REGION Network 6: setare bit 1 pentru SERVO6
   RUNG wire#powerrail
      I_Contact( "DB_HMI"."MAN/AUTO" )
      Contact( "DB_HMI_buttons"."ON/OFF_servo6" )
      wire#w1
      S_SR(operand := "DB_06_Write_Arduino".Servo6, r1 := wire#w3)
   END_RUNG
   RUNG wire#powerrail
      Contact( "DB_HMI"."MAN/AUTO" )
      Contact( "DB_Markers_Auto".servo6_auto )
   END_RUNG wire#w1
   RUNG wire#powerrail
      I_Contact( "DB_HMI"."MAN/AUTO" )
      I_Contact( "DB_HMI_buttons"."ON/OFF_servo6" )
      wire#w2
      R_Coil( "DB_HMI_buttons"."ON/OFF_servo6" )
   END_RUNG wire#w3
   RUNG wire#powerrail
      Contact( "DB_HMI"."MAN/AUTO" )
      I_Contact( "DB_Markers_Auto".servo6_auto )
   END_RUNG wire#w2
   RUNG wire#powerrail
      Contact( "DB_HMI_buttons".STOP )
   END_RUNG wire#w2
   // the same network as SCL:
   #_w1 := (NOT "DB_HMI"."MAN/AUTO" AND NOT "DB_HMI_buttons"."ON/OFF_servo6") OR ("DB_HMI"."MAN/AUTO" AND NOT "DB_Markers_Auto".servo6_auto) OR "DB_HMI_buttons".STOP;
   #_w2 := (NOT "DB_HMI"."MAN/AUTO" AND "DB_HMI_buttons"."ON/OFF_servo6") OR ("DB_HMI"."MAN/AUTO" AND "DB_Markers_Auto".servo6_auto);
   IF #_w1 THEN "DB_HMI_buttons"."ON/OFF_servo6" := FALSE; END_IF;
   IF #_w2 THEN
       "DB_06_Write_Arduino".Servo6 := TRUE;   // SR flip-flop
   END_IF;
   IF #_w1 THEN "DB_06_Write_Arduino".Servo6 := FALSE; END_IF;
END_REGION

REGION Network 7: setare bit stepper2_up
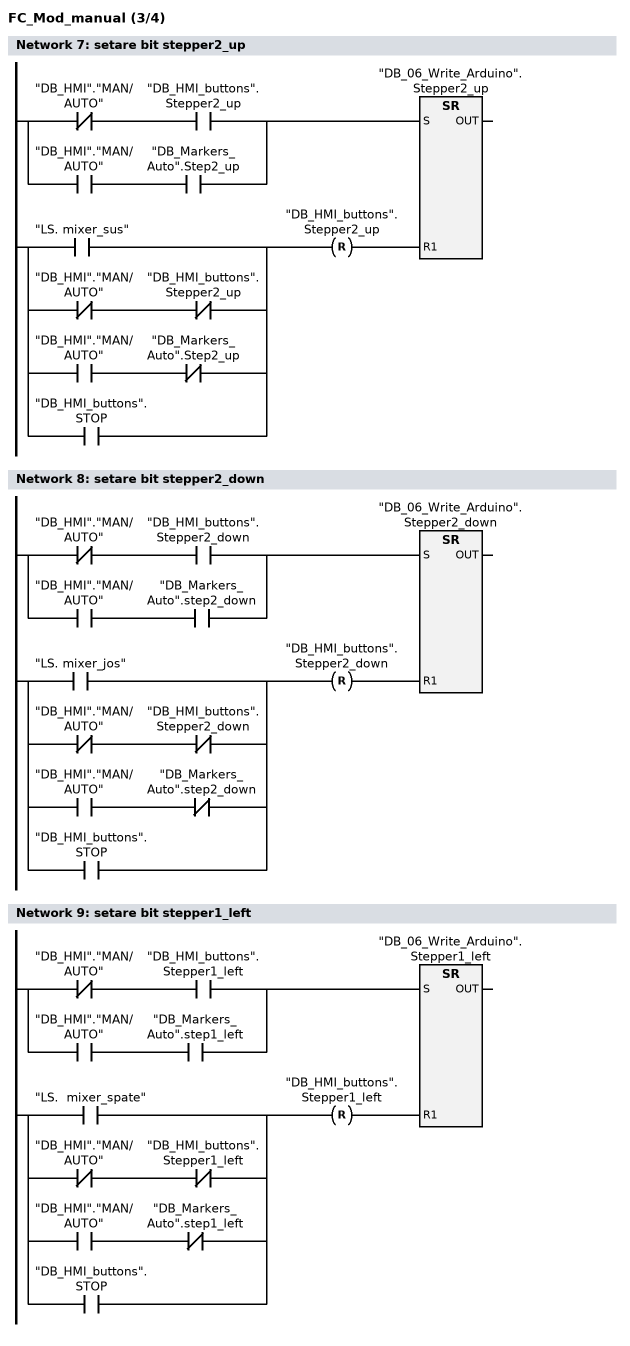
   RUNG wire#powerrail
      I_Contact( "DB_HMI"."MAN/AUTO" )
      Contact( "DB_HMI_buttons".Stepper2_up )
      wire#w1
      S_SR(operand := "DB_06_Write_Arduino".Stepper2_up, r1 := wire#w3)
   END_RUNG
   RUNG wire#powerrail
      Contact( "DB_HMI"."MAN/AUTO" )
      Contact( "DB_Markers_Auto".Step2_up )
   END_RUNG wire#w1
   RUNG wire#powerrail
      Contact( "LS. mixer_sus" )
      wire#w2
      R_Coil( "DB_HMI_buttons".Stepper2_up )
   END_RUNG wire#w3
   RUNG wire#powerrail
      I_Contact( "DB_HMI"."MAN/AUTO" )
      I_Contact( "DB_HMI_buttons".Stepper2_up )
   END_RUNG wire#w2
   RUNG wire#powerrail
      Contact( "DB_HMI"."MAN/AUTO" )
      I_Contact( "DB_Markers_Auto".Step2_up )
   END_RUNG wire#w2
   RUNG wire#powerrail
      Contact( "DB_HMI_buttons".STOP )
   END_RUNG wire#w2
   // the same network as SCL:
   #_w1 := "LS. mixer_sus" OR (NOT "DB_HMI"."MAN/AUTO" AND NOT "DB_HMI_buttons".Stepper2_up) OR ("DB_HMI"."MAN/AUTO" AND NOT "DB_Markers_Auto".Step2_up) OR "DB_HMI_buttons".STOP;
   #_w2 := (NOT "DB_HMI"."MAN/AUTO" AND "DB_HMI_buttons".Stepper2_up) OR ("DB_HMI"."MAN/AUTO" AND "DB_Markers_Auto".Step2_up);
   IF #_w1 THEN "DB_HMI_buttons".Stepper2_up := FALSE; END_IF;
   IF #_w2 THEN
       "DB_06_Write_Arduino".Stepper2_up := TRUE;   // SR flip-flop
   END_IF;
   IF #_w1 THEN "DB_06_Write_Arduino".Stepper2_up := FALSE; END_IF;
END_REGION

REGION Network 8: setare bit stepper2_down
   RUNG wire#powerrail
      I_Contact( "DB_HMI"."MAN/AUTO" )
      Contact( "DB_HMI_buttons".Stepper2_down )
      wire#w1
      S_SR(operand := "DB_06_Write_Arduino".Stepper2_down, r1 := wire#w3)
   END_RUNG
   RUNG wire#powerrail
      Contact( "DB_HMI"."MAN/AUTO" )
      Contact( "DB_Markers_Auto".step2_down )
   END_RUNG wire#w1
   RUNG wire#powerrail
      Contact( "LS. mixer_jos" )
      wire#w2
      R_Coil( "DB_HMI_buttons".Stepper2_down )
   END_RUNG wire#w3
   RUNG wire#powerrail
      I_Contact( "DB_HMI"."MAN/AUTO" )
      I_Contact( "DB_HMI_buttons".Stepper2_down )
   END_RUNG wire#w2
   RUNG wire#powerrail
      Contact( "DB_HMI"."MAN/AUTO" )
      I_Contact( "DB_Markers_Auto".step2_down )
   END_RUNG wire#w2
   RUNG wire#powerrail
      Contact( "DB_HMI_buttons".STOP )
   END_RUNG wire#w2
   // the same network as SCL:
   #_w1 := "LS. mixer_jos" OR (NOT "DB_HMI"."MAN/AUTO" AND NOT "DB_HMI_buttons".Stepper2_down) OR ("DB_HMI"."MAN/AUTO" AND NOT "DB_Markers_Auto".step2_down) OR "DB_HMI_buttons".STOP;
   #_w2 := (NOT "DB_HMI"."MAN/AUTO" AND "DB_HMI_buttons".Stepper2_down) OR ("DB_HMI"."MAN/AUTO" AND "DB_Markers_Auto".step2_down);
   IF #_w1 THEN "DB_HMI_buttons".Stepper2_down := FALSE; END_IF;
   IF #_w2 THEN
       "DB_06_Write_Arduino".Stepper2_down := TRUE;   // SR flip-flop
   END_IF;
   IF #_w1 THEN "DB_06_Write_Arduino".Stepper2_down := FALSE; END_IF;
END_REGION

REGION Network 9: setare bit stepper1_left
   RUNG wire#powerrail
      I_Contact( "DB_HMI"."MAN/AUTO" )
      Contact( "DB_HMI_buttons".Stepper1_left )
      wire#w1
      S_SR(operand := "DB_06_Write_Arduino".Stepper1_left, r1 := wire#w3)
   END_RUNG
   RUNG wire#powerrail
      Contact( "DB_HMI"."MAN/AUTO" )
      Contact( "DB_Markers_Auto".step1_left )
   END_RUNG wire#w1
   RUNG wire#powerrail
      Contact( "LS.  mixer_spate" )
      wire#w2
      R_Coil( "DB_HMI_buttons".Stepper1_left )
   END_RUNG wire#w3
   RUNG wire#powerrail
      I_Contact( "DB_HMI"."MAN/AUTO" )
      I_Contact( "DB_HMI_buttons".Stepper1_left )
   END_RUNG wire#w2
   RUNG wire#powerrail
      Contact( "DB_HMI"."MAN/AUTO" )
      I_Contact( "DB_Markers_Auto".step1_left )
   END_RUNG wire#w2
   RUNG wire#powerrail
      Contact( "DB_HMI_buttons".STOP )
   END_RUNG wire#w2
   // the same network as SCL:
   #_w1 := "LS.  mixer_spate" OR (NOT "DB_HMI"."MAN/AUTO" AND NOT "DB_HMI_buttons".Stepper1_left) OR ("DB_HMI"."MAN/AUTO" AND NOT "DB_Markers_Auto".step1_left) OR "DB_HMI_buttons".STOP;
   #_w2 := (NOT "DB_HMI"."MAN/AUTO" AND "DB_HMI_buttons".Stepper1_left) OR ("DB_HMI"."MAN/AUTO" AND "DB_Markers_Auto".step1_left);
   IF #_w1 THEN "DB_HMI_buttons".Stepper1_left := FALSE; END_IF;
   IF #_w2 THEN
       "DB_06_Write_Arduino".Stepper1_left := TRUE;   // SR flip-flop
   END_IF;
   IF #_w1 THEN "DB_06_Write_Arduino".Stepper1_left := FALSE; END_IF;
END_REGION

REGION Network 10: setare bit stepper1_right
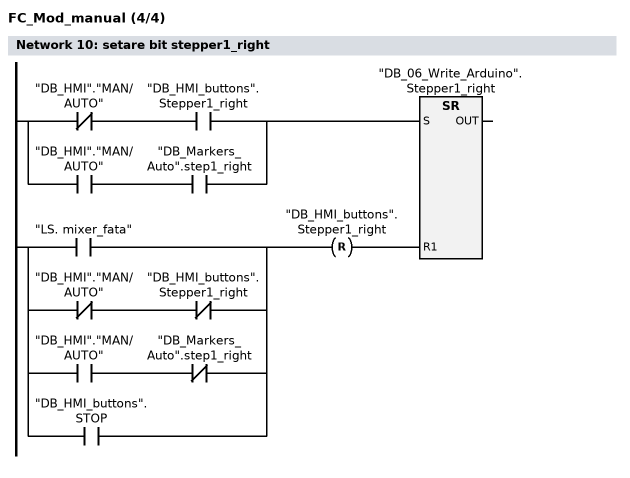
   RUNG wire#powerrail
      I_Contact( "DB_HMI"."MAN/AUTO" )
      Contact( "DB_HMI_buttons".Stepper1_right )
      wire#w1
      S_SR(operand := "DB_06_Write_Arduino".Stepper1_right, r1 := wire#w3)
   END_RUNG
   RUNG wire#powerrail
      Contact( "DB_HMI"."MAN/AUTO" )
      Contact( "DB_Markers_Auto".step1_right )
   END_RUNG wire#w1
   RUNG wire#powerrail
      Contact( "LS. mixer_fata" )
      wire#w2
      R_Coil( "DB_HMI_buttons".Stepper1_right )
   END_RUNG wire#w3
   RUNG wire#powerrail
      I_Contact( "DB_HMI"."MAN/AUTO" )
      I_Contact( "DB_HMI_buttons".Stepper1_right )
   END_RUNG wire#w2
   RUNG wire#powerrail
      Contact( "DB_HMI"."MAN/AUTO" )
      I_Contact( "DB_Markers_Auto".step1_right )
   END_RUNG wire#w2
   RUNG wire#powerrail
      Contact( "DB_HMI_buttons".STOP )
   END_RUNG wire#w2
   // the same network as SCL:
   #_w1 := "LS. mixer_fata" OR (NOT "DB_HMI"."MAN/AUTO" AND NOT "DB_HMI_buttons".Stepper1_right) OR ("DB_HMI"."MAN/AUTO" AND NOT "DB_Markers_Auto".step1_right) OR "DB_HMI_buttons".STOP;
   #_w2 := (NOT "DB_HMI"."MAN/AUTO" AND "DB_HMI_buttons".Stepper1_right) OR ("DB_HMI"."MAN/AUTO" AND "DB_Markers_Auto".step1_right);
   IF #_w1 THEN "DB_HMI_buttons".Stepper1_right := FALSE; END_IF;
   IF #_w2 THEN
       "DB_06_Write_Arduino".Stepper1_right := TRUE;   // SR flip-flop
   END_IF;
   IF #_w1 THEN "DB_06_Write_Arduino".Stepper1_right := FALSE; END_IF;
END_REGION
END_FUNCTION

FUNCTION "FC_select_reteta_FBD_language" : Void   // FC8, FBD
{ S7_Optimized_Access := 'TRUE' }
VERSION : 0.1
BEGIN

REGION Network 1: Reteta ciocolata neagra =1
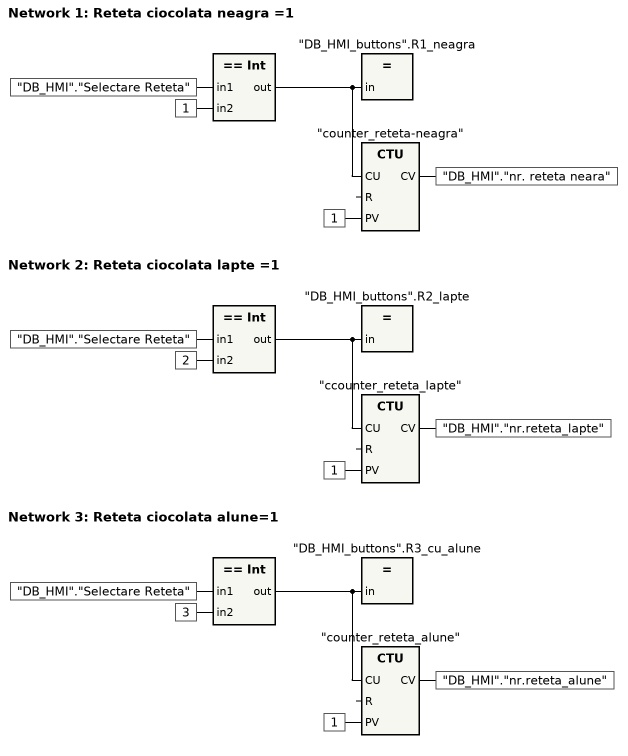
   "DB_HMI_buttons".R1_neagra := "DB_HMI"."Selectare Reteta" = 1;
   "counter_reteta-neagra".CTU(CU := "DB_HMI_buttons".R1_neagra, PV := 1, CV => "DB_HMI"."nr. reteta neara");
END_REGION

REGION Network 2: Reteta ciocolata lapte =1
   "DB_HMI_buttons".R2_lapte := "DB_HMI"."Selectare Reteta" = 2;
   "ccounter_reteta_lapte".CTU(CU := "DB_HMI_buttons".R2_lapte, PV := 1, CV => "DB_HMI"."nr.reteta_lapte");
END_REGION

REGION Network 3: Reteta ciocolata alune=1
   "DB_HMI_buttons".R3_cu_alune := "DB_HMI"."Selectare Reteta" = 3;
   "counter_reteta_alune".CTU(CU := "DB_HMI_buttons".R3_cu_alune, PV := 1, CV => "DB_HMI"."nr.reteta_alune");
END_REGION
END_FUNCTION

(* ===== HMI "HMI_RT_1" =====
system functions are stored by id; their names below are inferred from use
connection "Connection_1": ETHERNET, SMART_S7_1500_OMS
connection "HMI_Connection_1": ETHERNET, SMART_S7_1500_OMS

HMI tags "Default tag table"
   "LS_left" : Bool = PLC "LS.  mixer_spate" AT %I10.5, 1 s
   "LS_right" : Bool = PLC "LS. mixer_fata" AT %I10.2, 1 s
   "LS_up" : Bool = PLC "LS. mixer_sus" AT %I10.6, 1 s
   "LS_down" : Bool = PLC "LS. mixer_jos" AT %I10.1, 1 s
   "DB_HMI_BUTTON_DEV1:PLITA" : Bool = PLC DB_HMI_buttons.ON/OFF_plita AT %DB1.DBX0.0, 1 s
   "DB_HMI_BUTTON_DEV2:Mixer" : Bool = PLC DB_HMI_buttons.ON/OFF_mixer AT %DB1.DBX0.0, 1 s
   "DB_HMI_BUTTON_DEV2:Pompa" : Bool = PLC DB_HMI_buttons.ON/OFF_pompa AT %DB1.DBX0.0, 1 s
   "Reset ciuperca" : Bool = PLC DB_HMI_buttons.Reset_ciuperca AT %DB1.DBX0.0, 1 s
   "DB_06_Write_Arduino_Servo1" : Bool = PLC DB_06_Write_Arduino.Servo1 AT %DB6.DBX0.0, 1 s
   "DB_06_Write_Arduino_Servo2" : Bool = PLC DB_06_Write_Arduino.Servo2 AT %DB6.DBX0.1, 1 s
   "DB_06_Write_Arduino_Servo3" : Bool = PLC DB_06_Write_Arduino.Servo3 AT %DB6.DBX0.2, 1 s
   "DB_06_Write_Arduino_Servo4" : Bool = PLC DB_06_Write_Arduino.Servo4 AT %DB6.DBX0.3, 1 s
   "DB_06_Write_Arduino_Servo5" : Bool = PLC DB_06_Write_Arduino.Servo5 AT %DB6.DBX0.4, 1 s
   "DB_06_Write_Arduino_Servo6" : Bool = PLC DB_06_Write_Arduino.Servo6 AT %DB6.DBX0.5, 1 s
   "DB_HMI_buttons_ON/OFF_servo1" : Bool = PLC DB_HMI_buttons.ON/OFF_servo1, 1 s
   "ON/OFF_Servo1_HMI" : Word = PLC "ON/OFF_Servo1_HMI" AT %MW2, 1 s
   "ON/OFF_servo2_HMI" : Word = PLC "ON/OFF_servo2_HMI" AT %MW4, 1 s
   "ON/OFF_SERVO3_HMI" : Word = PLC "ON/OFF_SERVO3_HMI" AT %MW6, 1 s
   "ON/OFF_SERVO4_HMI" : Word = PLC "ON/OFF_SERVO4_HMI" AT %MW14, 1 s
   "ON/OFF_SERVO5_HMI" : Word = PLC "ON/OFF_SERVO5_HMI" AT %MW16, 1 s
   "ON/OFF_SERVO6_HMI" : Word = PLC "ON/OFF_SERVO6_HMI" AT %MW18, 1 s
   "ON/OFF_servo1" : Bool = PLC "ON/OFF_servo1" AT %M1.4, 1 s
   "DB_HMI_buttons_ON/OFF_servo2" : Bool = PLC DB_HMI_buttons.ON/OFF_servo2, 1 s
   "DB_HMI_buttons_ON/OFF_servo3" : Bool = PLC DB_HMI_buttons.ON/OFF_servo3, 1 s
   "DB_HMI_buttons_ON/OFF_servo4" : Bool = PLC DB_HMI_buttons.ON/OFF_servo4, 1 s
   "DB_HMI_buttons_ON/OFF_servo5" : Bool = PLC DB_HMI_buttons.ON/OFF_servo5, 1 s
   "DB_HMI_buttons_ON/OFF_servo6" : Bool = PLC DB_HMI_buttons.ON/OFF_servo6, 1 s
   "DB_HMI_buttons_Reset" : Bool = PLC DB_HMI_buttons.Reset, 1 s
   "DB_HMI_buttons_STOP" : Bool = PLC DB_HMI_buttons.STOP, 1 s
   "Reteta" : Int = PLC DB_HMI_buttons.Reteta_text_list AT %DB1.DBX0.0, 1 s
   "Start_initializare" : Bool = PLC DB_HMI_buttons.Start/Stop_initializare, 1 s
   "Start_proces" : Bool = PLC DB_HMI_buttons.Start/Stop_proces_auto, 1 s
   "DB_03_Read_Arduino_temp_citita" : Real = PLC DB_03_Read_Arduino.temp_citita AT %DB3.DBD0, 1 s
   "DB_06_Write_Arduino_Stepper2_up" : Bool = PLC DB_06_Write_Arduino.Stepper2_up AT %DB6.DBX1.0, 1 s
   "DB_06_Write_Arduino_Stepper2_down" : Bool = PLC DB_06_Write_Arduino.Stepper2_down AT %DB6.DBX1.1, 1 s
   "DB_HMI_buttons_Curatare" : Bool = PLC DB_HMI_buttons.Curatare, 1 s
   "DB_HMI_MAN/AUTO" : Bool = PLC DB_HMI.MAN/AUTO, 1 s
   "DB_HMI_Selectare Reteta" : Int = PLC DB_HMI."Selectare Reteta", 1 s
   "DB_06_Write_Arduino_Stepper1_left" : Bool = PLC DB_06_Write_Arduino.Stepper1_left AT %DB6.DBX0.6, 1 s
   "DB_06_Write_Arduino_Stepper1_right" : Bool = PLC DB_06_Write_Arduino.Stepper1_right AT %DB6.DBX0.7, 1 s
   "DB_HMI_buttons_Stepper1_left" : Bool = PLC DB_HMI_buttons.Stepper1_left, 1 s
   "DB_HMI_buttons_Stepper1_right" : Bool = PLC DB_HMI_buttons.Stepper1_right, 1 s
   "DB_HMI_buttons_Stop_stepper2" : Bool = PLC DB_HMI_buttons.Stop_stepper2, 1 s
   "DB_HMI_buttons_Stepper2_up" : Bool = PLC DB_HMI_buttons.Stepper2_up, 1 s
   "DB_HMI_buttons_Stop_stepper1" : Bool = PLC DB_HMI_buttons.Stop_stepper1, 1 s
   "DB_HMI_buttons_Stepper2_down" : Bool = PLC DB_HMI_buttons.Stepper2_down, 1 s
   "DB_HMI_buttons_Stop_stepper3" : Bool = PLC DB_HMI_buttons.Stop_stepper3, 1 s
   "DB_HMI_buttons_Stepper3_unloading" : Bool = PLC DB_HMI_buttons.Stepper3_unloading, 1 s
   "DB_HMI_buttons_Stepper3_loading" : Bool = PLC DB_HMI_buttons.Stepper3_loading, 1 s
   "DB_HMI_buttons_Initiere proces" : Bool = PLC DB_HMI_buttons."Initiere proces", 1 s
   "DB_HMI_Nr-pas_auto" : Int = PLC DB_HMI.Nr-pas_auto, 1 s
   "DB_HMI_Bypass-pompa" : Bool = PLC DB_HMI.Bypass-pompa, 1 s
   "DB_HMI_bypass_plita" : Bool = PLC DB_HMI.bypass_plita, 1 s
   "DB_HMI_bypass_mixer" : Bool = PLC DB_HMI.bypass_mixer, 1 s
   "PLC_1_DB_HMI_buttons_R3_cu_alune" : Bool = PLC DB_HMI_buttons.R3_cu_alune, 1 s
   "PLC_1_DB_HMI_buttons_R2_lapte" : Bool = PLC DB_HMI_buttons.R2_lapte, 1 s
   "PLC_1_DB_HMI_buttons_R1_neagra" : Bool = PLC DB_HMI_buttons.R1_neagra, 1 s
   "PLC_1_DB_Markers_M_Auto" : Bool = PLC DB_Markers.M_Auto, 1 s
   "PLC_1_DB_Markers_M_Manual" : Bool = PLC DB_Markers.M_Manual, 1 s

HMI tags "Alarms"
   "Alarm_mod_manual" : Word = PLC DB_Messages.B002, 1 s
   "Alarm_mod_auto" : Word = PLC DB_Messages.B003 AT %DB1.DBW0, 1 s
   "Alarm_servo1_on" : Word = PLC DB_Messages.B009 AT %DB1.DBW0, 1 s
   "Alarm_stepper1_on" : Word = PLC DB_Messages.B011 AT %DB1.DBW0, 1 s
   "Alarm_stepper2-on" : Word = PLC DB_Messages.B012 AT %DB1.DBW0, 1 s
   "Alarm_stepper3-on" : Word = PLC DB_Messages.B013 AT %DB1.DBW0, 1 s
   "Alarm bol in poz necoresp" : Word = PLC DB_Messages.B006 AT %DB1.DBW0, 1 s
   "Alarm_plita on" : Word = PLC DB_Messages.B008 AT %DB1.DBW0, 1 s
   "Alarm_mixer_poz_necoresp" : Word = PLC DB_Messages.B005 AT %DB1.DBW0, 1 s

discrete alarms
   1: 'Statia e in modul manual!', class InfoMessages, trigger "Alarm_mod_manual" bit 0
   2: 'Statia este in modul automat!', class InfoMessages, trigger "Alarm_mod_auto" bit 0
   3: 'Valva1 e deschisa!', class InfoMessages, trigger "Alarm_servo1_on" bit 0
   4: 'Mixerul se deplaseaza pe orizontala.', class InfoMessages, trigger "Alarm_stepper1_on" bit 0
   5: 'Mixerul se deplaseaza pe verticala', class InfoMessages, trigger "Alarm_stepper2-on" bit 0
   6: 'Bolul de amestec este in proces de basculare/revenire.', class InfoMessages, trigger "Alarm_stepper3-on" bit 0
   7: 'Mixerul se afla intr-o pozitie necorespunzatoare!', class Warnings, trigger "Alarm_mixer_poz_necoresp" bit 0

text list "Retete": 0 'Selectare reteta'; 1 'Ciocolata neagra'; 2 'Ciocolata cu lapte'; 3 'Ciocolata cu alune'

Template "Template_1" 800x480
   Button "Exit" at 714,429 size 71x50; TextOff 'Exit'; PictureOff "ExitRuntime_KTP700_Basic_PN_TR"; PictureOn "ExitRuntime_KTP700_Basic_PN_TR"
      on Release: StopRuntime(0)
   Button "Template_Button" at 614,429 size 71x50; TextOff 'Text'
   Button "Template_Button_1" at 516,429 size 71x50; TextOff 'Text'
   Button "Template_Button_2" at 379,429 size 71x50; TextOff 'Text'
   Button "Template_Button_3" at 293,429 size 71x50; TextOff 'Dozare'
   Button "Template_Button_4" at 112,429 size 158x50; TextOff 'Pornire motoare'
   Button "Start screen" at 14,429 size 71x50; TextOff 'Start screen'; PictureOff "NavigateHome_KTP700_Basic_PN_TR"; PictureOn "NavigateHome_KTP700_Basic_PN_TR"
      on Release: ActivateScreen("Screen 1", 0)
   GraphicView "Logo" at 0,0 size 91x51; Picture "Logo of HMI_1"

screen "Screen 1" 800x480
   TextField "Text field_1" at 171,231 size 583x47; Text 'LINIE AUTOMATA SI MANUALA'
   Button "Button_1" at 11,172 size 132x64; TextOff 'Testare in mod manual'
      on Press: ActivateScreen("MANUAL", 0)
      Visibility <- "DB_HMI_MAN/AUTO"
   GraphicView "Graphic view_2" at 549,78 size 233x178; Picture "—Pngtree—cartoon hand drawn minimalistic splash_1"
   TextField "Text field_2" at 244,278 size 465x39; Text 'DE FABRICATIE A CIOCOLATEI'
   Button "Button_2" at 11,172 size 132x64; TextOff 'Mod automat'
      on Press: ActivateScreen("Automat", 0)
      Visibility <- "DB_HMI_MAN/AUTO"
   Switch "Switch_1" at 11,101 size 132x64; CaptionText 'Switch'; TextOff 'Manual'; TextOn 'Auto'
      ProcessValue <- "DB_HMI_MAN/AUTO"
      Appearance <- "DB_HMI_MAN/AUTO"
   Circle "Circle_5" at 150,115 size 21x21
      Appearance <- "DB_HMI_MAN/AUTO"
   Button "Button_5" at 656,409 size 144x71; TextOff 'Inchide'
      on Press: StopRuntime(0)
   GraphicView "Graphic view_1" at 8,4 size 177x37; Picture "Siemens_AG_logo.svg"
   GraphicView "Graphic view_3" at 98,251 size 233x178; Picture "—Pngtree—cartoon hand drawn minimalistic splash_1"
   TextField "Text field_3" at 11,75 size 202x23; Text 'Selectati modul de lucru'
   Button "Button_6" at 18,413 size 146x67; TextOff 'Parametri'
      on Press: ActivateScreen("Parametri", 0)
   DateTimeField "Date/time field_1" at 576,9 size 219x32
   Button "Button_7" at 189,413 size 146x67; TextOff 'Mesaje/Erori'
      on Press: ActivateScreen("Mesaje/Erori", 0)
   GraphicView "Graphic view_4" at 758,423 size 42x43; Picture "Graphic_47"
   TextField "Text field_8" at 435,52 size 245x23; Text 'Statia functioneaza in modul:'
   TextField "Text field_10" at 555,75 size 88x27; Text 'MANUAL'
      Visibility <- "DB_HMI_MAN/AUTO"
   TextField "Text field_9" at 538,75 size 101x27; Text 'AUTOMAT'
      Visibility <- "DB_HMI_MAN/AUTO"
   Ellipse "Ellipse_2" at 642,77 size 25x24
      Appearance <- "DB_HMI_MAN/AUTO"
      Visibility <- "DB_HMI_MAN/AUTO"
   Ellipse "Ellipse_1" at 642,76 size 25x24
      Visibility <- "DB_HMI_MAN/AUTO"
      Appearance <- "DB_HMI_MAN/AUTO"
   Button "Button_3" at 691,52 size 102x49; TextOff 'Stop'
      on Press: SetBit("DB_HMI_buttons_STOP")
      Visibility <- "DB_HMI_buttons_STOP"
   Button "Button_4" at 691,53 size 102x49; TextOff 'Resetare'
      on Press: ResetBit("DB_HMI_buttons_STOP")
      Visibility <- "DB_HMI_buttons_STOP"
      Appearance <- "DB_HMI_buttons_STOP"

screen "MANUAL" 800x480
   Button "Button_2" at 399,173 size 165x78; TextOff 'Mixare'
      on Click: ActivateScreen("MIXARE", 0)
   Button "Button_1" at 211,173 size 165x78; TextOff 'Dozare'
      on Click: ActivateScreen("DOZARE", 0)
   Button "Button_3" at 211,278 size 165x78; TextOff 'Topire'
      on Click: ActivateScreen("Pornire plita", 0)
   Button "Button_4" at 399,278 size 165x79; TextOff 'Adaugare apa'
      on Click: ActivateScreen("pornire pompa", 0)
   Button "Button_13" at 654,413 size 146x67; TextOff 'Inapoi'
      on Click: ActivateScreen("Screen 1", 0)
   Button "Button_5" at 693,56 size 102x49; TextOff 'Stop'
      on Press: SetBit("DB_HMI_buttons_STOP")
      Visibility <- "DB_HMI_buttons_STOP"
   Button "Button_6" at 693,56 size 102x49; TextOff 'Resetare'
      on Press: ResetBit("DB_HMI_buttons_STOP")
      Visibility <- "DB_HMI_buttons_STOP"
      Appearance <- "DB_HMI_buttons_STOP"
   TextField "Text field_1" at 229,84 size 306x34; Text 'Testare in mod MANUAL'
   GraphicView "Graphic view_1" at 8,4 size 177x37; Picture "Siemens_AG_logo.svg"
   DateTimeField "Date/time field_1" at 576,9 size 219x32
   Button "Button_8" at 20,413 size 146x67; TextOff 'Parametri'
      on Press: ActivateScreen("Parametri", 0)
   Button "Button_7" at 184,413 size 146x67; TextOff 'Mesaje/Erori'
      on Press: ActivateScreen("Mesaje/Erori", 0)

screen "DOZARE" 800x480
   GraphicView "Graphic view_1" at 141,130 size 155x135; Picture "Graphic_1"
   GraphicView "Graphic view_2" at 209,242 size 25x199; Picture "Graphic_16"
   Group "Group" at 141,130 size 155x311; Picture "Graphic_1"
   GraphicView "Graphic view_7" at 200,241 size 39x24; Picture "Graphic_28"
   GraphicView "Graphic view_8" at 197,355 size 42x27; Picture "Graphic_28"
   Group "Group_1" at 141,130 size 155x311; Picture "Graphic_1"
   Group "Group_3" at 363,130 size 155x311; Picture "Graphic_1"
   Group "Group_5" at 591,131 size 155x311; Picture "Graphic_1"
   Button "Button_1" at 86,233 size 96x45; TextOff 'ON/OFF Servo1'
      on Press: InvertBit("DB_HMI_buttons_ON/OFF_servo1")
   Button "Button_7" at 85,345 size 96x45; TextOff 'ON/OFF Servo4'
      on Press: InvertBit("DB_HMI_buttons_ON/OFF_servo4")
   Button "Button_2" at 309,232 size 96x45; TextOff 'ON/OFF Servo2'
      on Press: InvertBit("DB_HMI_buttons_ON/OFF_servo2")
   Button "Button_3" at 309,343 size 96x45; TextOff 'ON/OFF Servo5'
      on Press: InvertBit("DB_HMI_buttons_ON/OFF_servo5")
   Button "Button_4" at 539,233 size 96x45; TextOff 'ON/OFF Servo3'
      on Press: InvertBit("DB_HMI_buttons_ON/OFF_servo3")
   Button "Button_5" at 536,343 size 96x45; TextOff 'ON/OFF Servo6'
      on Press: InvertBit("DB_HMI_buttons_ON/OFF_servo6")
   Circle "Circle_1" at 58,243 size 21x21
      Appearance <- "DB_HMI_buttons_ON/OFF_servo1"
   Circle "Circle_2" at 58,353 size 21x21
      Visibility <- "ON/OFF_servo2_HMI"
      Appearance <- "DB_HMI_buttons_ON/OFF_servo4"
   Circle "Circle_3" at 278,239 size 21x21
      Visibility <- "ON/OFF_SERVO3_HMI"
      Appearance <- "DB_HMI_buttons_ON/OFF_servo2"
   Circle "Circle_4" at 278,353 size 21x21
      Visibility <- "ON/OFF_SERVO4_HMI"
      Appearance <- "DB_HMI_buttons_ON/OFF_servo5"
   Circle "Circle_5" at 505,244 size 21x21
      Visibility <- "ON/OFF_SERVO5_HMI"
      Appearance <- "DB_HMI_buttons_ON/OFF_servo3"
   Circle "Circle_6" at 505,352 size 21x21
      Visibility <- "ON/OFF_SERVO6_HMI"
      Appearance <- "DB_HMI_buttons_ON/OFF_servo6"
   TextField "Text field_1" at 244,54 size 295x34; Text 'Dozarea ingredientelor'
   Button "Button_6" at 693,46 size 102x49; TextOff 'Stop'
      on Press: SetBit("DB_HMI_buttons_STOP")
      Visibility <- "DB_HMI_buttons_STOP"
   Button "Button_8" at 692,46 size 102x49; TextOff 'Resetare'
      on Press: ResetBit("DB_HMI_buttons_STOP")
      Visibility <- "DB_HMI_buttons_STOP"
      Appearance <- "DB_HMI_buttons_STOP"
   GraphicView "Graphic view_13" at 8,4 size 177x37; Picture "Siemens_AG_logo.svg"
   DateTimeField "Date/time field_1" at 576,9 size 219x32
   Button "Button_13" at 654,413 size 146x67; TextOff 'Inapoi'
      on Click: ActivateScreen("MANUAL", 0)
   GraphicView "Graphic view_3" at 363,130 size 155x135; Picture "Graphic_1"
   GraphicView "Graphic view_4" at 431,242 size 25x199; Picture "Graphic_16"
   Group "Group_2" at 363,130 size 155x311; Picture "Graphic_1"
   GraphicView "Graphic view_5" at 422,241 size 39x24; Picture "Graphic_28"
   GraphicView "Graphic view_6" at 419,355 size 42x27; Picture "Graphic_28"
   GraphicView "Graphic view_9" at 591,131 size 155x135; Picture "Graphic_1"
   GraphicView "Graphic view_10" at 659,243 size 25x199; Picture "Graphic_16"
   Group "Group_4" at 591,131 size 155x311; Picture "Graphic_1"
   GraphicView "Graphic view_11" at 650,242 size 39x24; Picture "Graphic_28"
   GraphicView "Graphic view_12" at 647,356 size 42x27; Picture "Graphic_28"

screen "Pornire plita" 800x480
   GraphicView "Graphic view_1" at 328,229 size 113x133; Picture "189956"
   Button "Button_1" at 318,367 size 130x70; TextOff 'Plita ON/OFF'
      on Press: InvertBit("DB_HMI_BUTTON_DEV1:PLITA")
      Appearance <- "DB_HMI_BUTTON_DEV1:PLITA"
   TextField "Text field_1" at 267,80 size 204x34; Text 'Topire ciocolata'
   Button "Button_13" at 654,413 size 146x67; TextOff 'Inapoi'
      on Click: ActivateScreen("MANUAL", 0)
   GraphicView "Graphic view_13" at 8,4 size 177x37; Picture "Siemens_AG_logo.svg"
   DateTimeField "Date/time field_1" at 576,9 size 219x32
   Button "Button_2" at 693,46 size 102x49; TextOff 'Stop'
      on Press: SetBit("DB_HMI_buttons_STOP")
      Visibility <- "DB_HMI_buttons_STOP"
   Button "Button_4" at 692,46 size 102x49; TextOff 'Resetare'
      on Press: ResetBit("DB_HMI_buttons_STOP")
      Visibility <- "DB_HMI_buttons_STOP"
      Appearance <- "DB_HMI_buttons_STOP"
   AlarmView "Alarm view_1" at 16,128 size 769x101; ColumnTextAlarmText 'Mesaje/Erori'
   Circle "Circle_1" at 286,392 size 21x21
      Appearance <- "DB_HMI_BUTTON_DEV1:PLITA"

screen "MIXARE" 800x480
   GraphicView "Graphic view_1" at 94,153 size 265x222; Picture "Graphic_14"
   TextField "Text field_1" at 162,89 size 439x34; Text 'Setati mixerul in pozitia de mixare'
   Circle "Circle_1" at 135,336 size 21x21
      Appearance <- "DB_HMI_BUTTON_DEV2:Mixer"
   Button "Button_13" at 654,413 size 146x67; TextOff 'Inapoi'
      on Click: ActivateScreen("MANUAL", 0)
   GraphicView "Graphic view_13" at 8,4 size 177x37; Picture "Siemens_AG_logo.svg"
   Button "Button_2" at 693,46 size 102x49; TextOff 'Stop'
      on Press: SetBit("DB_HMI_buttons_STOP")
      Visibility <- "DB_HMI_buttons_STOP"
   Button "Button_4" at 693,46 size 102x49; TextOff 'Resetare'
      on Press: ResetBit("DB_HMI_buttons_STOP")
      Visibility <- "DB_HMI_buttons_STOP"
      Appearance <- "DB_HMI_buttons_STOP"
   DateTimeField "Date/time field_1" at 576,9 size 219x32
   Button "Button_7" at 364,189 size 102x49; TextOff 'Sus ON/OFF'
      on Press: SetBit("DB_HMI_buttons_Stepper2_up")
      Appearance <- "DB_06_Write_Arduino_Stepper2_up"
   Button "Button_3" at 552,189 size 102x49; TextOff 'Stanga ON/OFF'
      Appearance <- "DB_06_Write_Arduino_Stepper1_left"
      on Press: SetBit("DB_HMI_buttons_Stepper1_left")
   Button "Button_5" at 364,275 size 102x49; TextOff 'Jos ON/OFF'
      Appearance <- "DB_06_Write_Arduino_Stepper2_down"
      on Press: SetBit("DB_HMI_buttons_Stepper2_down")
   Button "Button_6" at 556,275 size 102x49; TextOff 'Dreapta ON/OFF'
      on Press: SetBit("DB_HMI_buttons_Stepper1_right")
      Appearance <- "DB_06_Write_Arduino_Stepper1_right"
   Button "Button_1" at 162,324 size 102x49; TextOff 'ON/OFF'
      on Press: InvertBit("DB_HMI_BUTTON_DEV2:Mixer")
      Appearance <- "DB_HMI_BUTTON_DEV2:Mixer"

screen "pornire pompa" 800x480
   TextField "Text field_1" at 301,57 size 179x34; Text 'Adaugare apa'
   DateTimeField "Date/time field_1" at 576,9 size 219x32
   GraphicView "Graphic view_13" at 8,4 size 177x37; Picture "Siemens_AG_logo.svg"
   Button "Button_3" at 693,46 size 102x49; TextOff 'Stop'
      on Press: SetBit("DB_HMI_buttons_STOP")
      Visibility <- "DB_HMI_buttons_STOP"
   Button "Button_4" at 692,46 size 102x49; TextOff 'Resetare'
      on Press: ResetBit("DB_HMI_buttons_STOP")
      Visibility <- "DB_HMI_buttons_STOP"
      Appearance <- "DB_HMI_buttons_STOP"
   Button "Button_13" at 654,413 size 146x67; TextOff 'Inapoi'
      on Press: ActivateScreen("MANUAL", 0)
   AlarmView "Alarm view_1" at 23,111 size 768x101; ColumnTextAlarmText 'Mesaje/Erori'
   Button "Button_1" at 333,349 size 130x70; TextOff 'Pompa ON/OFF'
      on Press: InvertBit("DB_HMI_BUTTON_DEV2:Pompa")
      Appearance <- "DB_HMI_BUTTON_DEV2:Pompa"
   GraphicView "Graphic view_2" at 343,213 size 141x169; Picture "Graphic_29"
   Circle "Circle_1" at 298,373 size 21x21
      Appearance <- "DB_HMI_BUTTON_DEV2:Pompa"

screen "Automat" 800x480
   Button "Button_13" at 654,413 size 146x67; TextOff 'Inapoi'
      on Press: ActivateScreen("Screen 1", 0)
   Button "Button_4" at 234,283 size 102x49; TextOff 'Start/Stop proces'
      on Press: SetBit("Start_proces")
      on Release: ResetBit("Start_proces")
      Appearance <- "Start_proces"
   TextField "Text field_1" at 673,186 size 118x23; Text 'Temperatura:'
   SymbolicIOField "Symbolic I/O field_1" at 255,107 size 284x37; TextOff '0'; TextOn '1'; TextList "Retete"
      TextList <- "Reteta"
      ProcessValue <- "DB_HMI_Selectare Reteta"
   TextField "Text field_2" at 292,66 size 195x34; Text 'Mod AUTOMAT'
   Button "Button_1" at 234,357 size 102x49; TextOff 'Start/Stop curatare'
      on Press: SetBit("DB_HMI_buttons_Curatare")
      on Release: ResetBit("DB_HMI_buttons_Curatare")
      Appearance <- "DB_HMI_buttons_Curatare"
   Button "Button_3" at 689,56 size 102x49; TextOff 'Stop'
      on Press: SetBit("DB_HMI_buttons_STOP")
      Visibility <- "DB_HMI_buttons_STOP"
   Button "Button_5" at 689,56 size 102x49; TextOff 'Resetare'
      on Press: ResetBit("DB_HMI_buttons_STOP")
      Visibility <- "DB_HMI_buttons_STOP"
      Appearance <- "DB_HMI_buttons_STOP"
   Button "Button_2" at 147,204 size 102x49; TextOff 'Initiere proces'
      on Press: SetBit("DB_HMI_buttons_Initiere proces")
      on Release: ResetBit("DB_HMI_buttons_Initiere proces")
      Appearance <- "DB_HMI_buttons_Initiere proces"
   IOField "I/O field_3" at 731,136 size 65x34; FormatPattern 999
      ProcessValue <- "DB_HMI_Nr-pas_auto"
   TextField "Text field_3" at 656,141 size 73x23; Text 'Nr. pas :'
   GraphicView "Graphic view_1" at 2,0 size 177x37; Picture "Siemens_AG_logo.svg"
   DateTimeField "Date/time field_1" at 576,9 size 219x32
   Button "Button_6" at 18,424 size 102x49; TextOff 'Bypass pompa'
      on Press: SetBit("DB_HMI_Bypass-pompa")
      on Release: ResetBit("DB_HMI_Bypass-pompa")
   Button "Button_7" at 136,424 size 102x49; TextOff 'Bypass plita'
      on Release: ResetBit("DB_HMI_bypass_plita")
      on Press: SetBit("DB_HMI_bypass_plita")
   Button "Button_8" at 255,424 size 102x49; TextOff 'Bypass mixer'
      on Release: ResetBit("DB_HMI_bypass_mixer")
      on Press: SetBit("DB_HMI_bypass_mixer")
   IOField "I/O field_2" at 695,209 size 96x32; FormatPattern s999.999
      ProcessValue <- "DB_03_Read_Arduino_temp_citita"
   TextField "Text field_4" at 211,151 size 192x23; Text 'Reteta selectata este:'
   TextField "Text field_5" at 405,151 size 154x23; Text 'Ciocolata cu alune'
      Visibility <- "PLC_1_DB_HMI_buttons_R3_cu_alune"
   TextField "Text field_6" at 405,151 size 151x23; Text 'Ciocolata cu lapte'
      Visibility <- "PLC_1_DB_HMI_buttons_R2_lapte"
   TextField "Text field_7" at 405,151 size 143x23; Text 'Ciocolata neagra'
      Visibility <- "PLC_1_DB_HMI_buttons_R1_neagra"
   TextField "Text field_8" at 10,56 size 245x23; Text 'Statia functioneaza in modul:'
   TextField "Text field_9" at 19,77 size 101x27; Text 'AUTOMAT'
      Visibility <- "DB_HMI_MAN/AUTO"
   Ellipse "Ellipse_1" at 123,77 size 25x24
      Appearance <- "DB_HMI_MAN/AUTO"
      Visibility <- "DB_HMI_MAN/AUTO"
   TextField "Text field_10" at 30,76 size 88x27; Text 'MANUAL'
      Visibility <- "DB_HMI_MAN/AUTO"
   Ellipse "Ellipse_2" at 123,78 size 25x24
      Visibility <- "DB_HMI_MAN/AUTO"
      Appearance <- "DB_HMI_MAN/AUTO"
   TextField "Text field_11" at 10,204 size 129x42; Text 'Initiere proces in asteptare:'
      Visibility <- "DB_HMI_buttons_Initiere proces"
   TextField "Text field_13" at 10,205 size 130x42; Text 'Procesul a fost initiat!'
      Visibility <- "DB_HMI_buttons_Initiere proces"
   TextField "Text field_12" at 11,281 size 203x61; Text 'Dupa selectarea retetei apasati butonul pentru a porni procesul:'
      Visibility <- "Start_proces"
   TextField "Text field_14" at 50,297 size 159x23; Text 'Procesul a inceput!'
      Visibility <- "Start_proces"
   TextField "Text field_15" at 8,357 size 226x42; Text 'Pentru a curata vasul de amestec, selectati butonul:'
      Visibility <- "DB_HMI_buttons_Curatare"
   TextField "Text field_16" at 5,369 size 226x23; Text 'Ciclu de curatare in proces!'
      Visibility <- "DB_HMI_buttons_Curatare"

screen "Parametri" 800x480
   GraphicView "Graphic view_13" at 8,4 size 177x37; Picture "Siemens_AG_logo.svg"
   DateTimeField "Date/time field_1" at 576,9 size 219x32
   TextField "Text field_1" at 293,69 size 213x34; Text 'Parametri retete'
   TextField "Text field_2" at 95,127 size 151x23; Text 'Ciocolata cu lapte'
   TextField "Text field_3" at 304,127 size 154x23; Text 'Ciocolata cu alune'
   TextField "Text field_4" at 534,127 size 143x23; Text 'Ciocolata neagra'
   TextField "Text field_5" at 82,166 size 160x44; Text 'Timpi pentru dozare:'
   TextField "Text field_6" at 82,196 size 93x80; Text '- valva 1: 5s - valva 2: 5s - valva 4: 5s - valva 5: 5s'
   TextField "Text field_7" at 287,196 size 93x80; Text '- valva 1: 5s - valva 2: 7s - valva 4: 5s - valva 5: 7s'
   TextField "Text field_8" at 282,166 size 160x44; Text 'Timpi pentru dozare:'
   TextField "Text field_9" at 520,166 size 160x44; Text 'Timpi pentru dozare:'
   TextField "Text field_10" at 520,196 size 93x80; Text '- valva 1: 6s - valva 2: 6s - valva 4: 5s - valva 5: 5s'
   TextField "Text field_11" at 77,276 size 161x44; Text 'Timpi pentru mixare:'
   TextField "Text field_12" at 282,275 size 161x44; Text 'Timpi pentru mixare:'
   TextField "Text field_13" at 516,278 size 161x44; Text 'Timpi pentru mixare:'
   TextField "Text field_14" at 83,297 size 32x23; Text '- 5s'
   TextField "Text field_15" at 272,299 size 32x23; Text '- 5s'
   TextField "Text field_16" at 520,301 size 32x23; Text '- 5s'
   TextField "Text field_17" at 76,323 size 170x44; Text 'Timpi pentru incalzire:'
   TextField "Text field_18" at 280,321 size 170x44; Text 'Timpi pentru incalzire:'
   TextField "Text field_19" at 518,321 size 170x44; Text 'Timpi pentru incalzire:'
   TextField "Text field_20" at 83,346 size 32x23; Text '- 7s'
   TextField "Text field_22" at 272,343 size 41x23; Text '- 10s'
   TextField "Text field_23" at 520,342 size 41x23; Text '- 15s'
   Button "Button_13" at 657,423 size 143x57; TextOff 'Inapoi'
      on Click: ActivateScreen("Screen 1", 0)
   TextField "Text field_21" at 75,374 size 107x24; Text 'Temperatura:'
   TextField "Text field_24" at 280,375 size 107x24; Text 'Temperatura:'
   TextField "Text field_25" at 519,376 size 107x24; Text 'Temperatura:'
   TextField "Text field_26" at 84,394 size 142x23; Text '- 100 grade Celsius'
   TextField "Text field_27" at 269,394 size 142x23; Text '- 150 grade Celsius'
   TextField "Text field_28" at 515,394 size 142x23; Text '- 130 grade Celsius'

screen "Mesaje/Erori" 800x480
   GraphicView "Graphic view_1" at 8,4 size 177x37; Picture "Siemens_AG_logo.svg"
   DateTimeField "Date/time field_1" at 576,9 size 219x32
   TextField "Text field_1" at 301,67 size 168x34; Text 'Mesaje/Erori'
   AlarmView "Alarm view_1" at 23,123 size 759x273; ColumnTextAlarmText 'Mesaje/Erori'
   Button "Button_13" at 654,413 size 146x67; TextOff 'Inapoi'
      on Click: ActivateScreen("Screen 1", 0)
*)